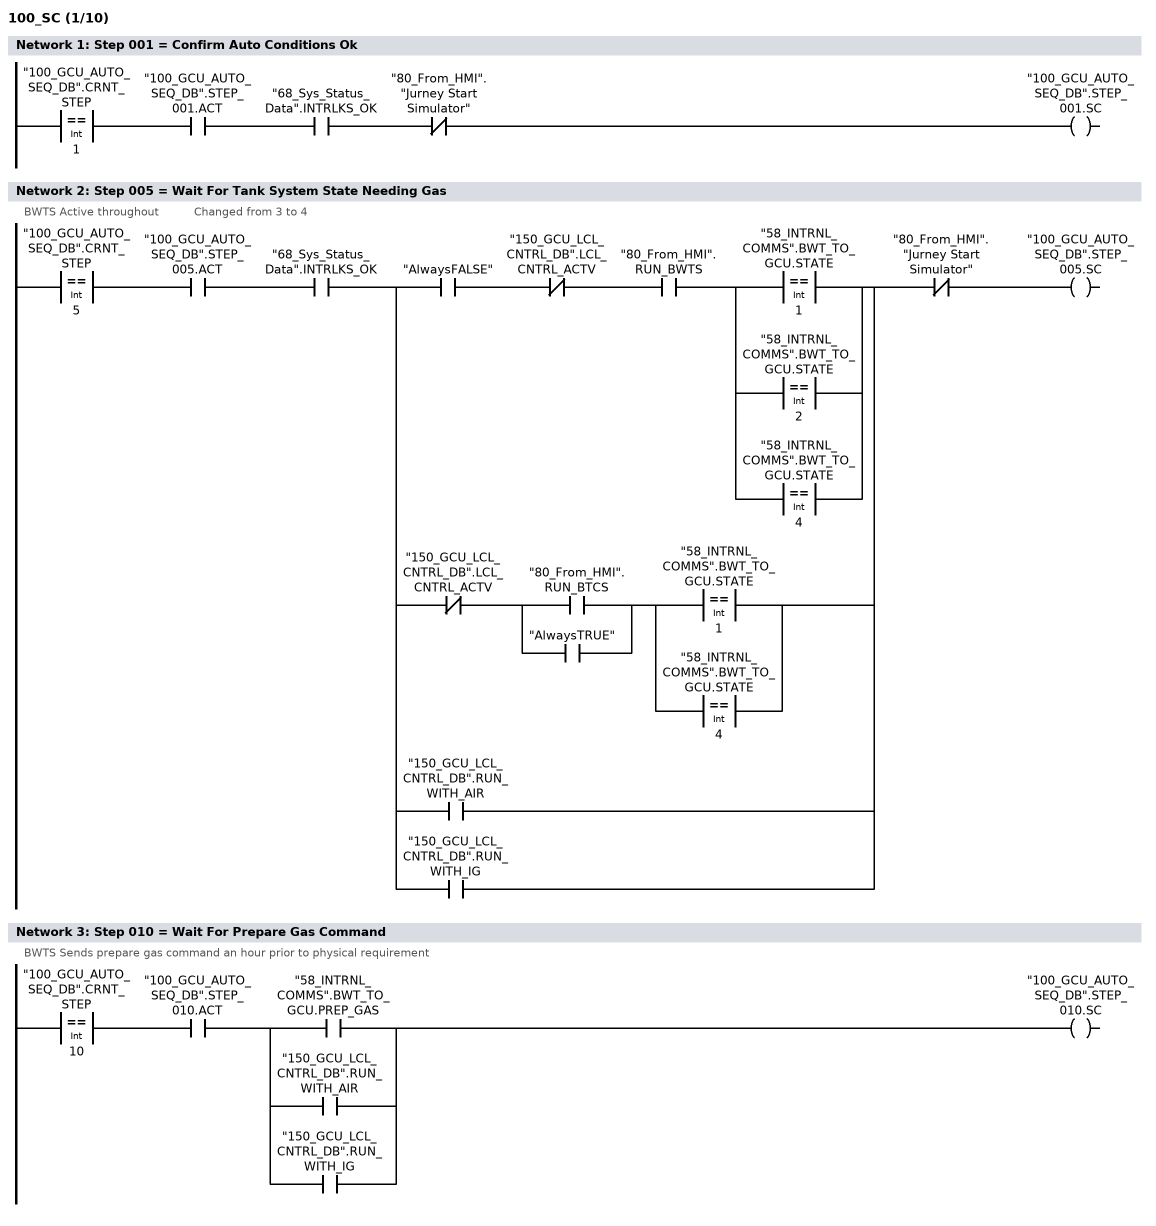
   RUNG wire#powerrail
      { S7_Templates := "SrcType := Int" } EQ_Contact(in1 := "100_GCU_AUTO_SEQ_DB".CRNT_STEP, in2 := 1)
      Contact( "100_GCU_AUTO_SEQ_DB".STEP_001.ACT )
      Contact( "68_Sys_Status_Data".INTRLKS_OK )
      I_Contact( "80_From_HMI"."Jurney Start Simulator" )
      Coil( "100_GCU_AUTO_SEQ_DB".STEP_001.SC )
   END_RUNG
   // the same network as SCL:
   "100_GCU_AUTO_SEQ_DB".STEP_001.SC := ("100_GCU_AUTO_SEQ_DB".CRNT_STEP = 1) AND "100_GCU_AUTO_SEQ_DB".STEP_001.ACT AND "68_Sys_Status_Data".INTRLKS_OK AND NOT "80_From_HMI"."Jurney Start Simulator";
END_REGION

REGION Network 2: Step 005 = Wait For Tank System State Needing Gas
   // BWTS Active throughout          Changed from 3 to 4
   RUNG wire#powerrail
      { S7_Templates := "SrcType := Int" } EQ_Contact(in1 := "100_GCU_AUTO_SEQ_DB".CRNT_STEP, in2 := 5)
      Contact( "100_GCU_AUTO_SEQ_DB".STEP_005.ACT )
      Contact( "68_Sys_Status_Data".INTRLKS_OK )
      wire#w1
      Contact( "AlwaysFALSE" )
      I_Contact( "150_GCU_LCL_CNTRL_DB".LCL_CNTRL_ACTV )
      Contact( "80_From_HMI".RUN_BWTS )
      wire#w2
      { S7_Templates := "SrcType := Int" } EQ_Contact(in1 := "58_INTRNL_COMMS".BWT_TO_GCU.STATE, in2 := 1)
      wire#w3
      I_Contact( "80_From_HMI"."Jurney Start Simulator" )
      Coil( "100_GCU_AUTO_SEQ_DB".STEP_005.SC )
   END_RUNG
   RUNG wire#w2
      { S7_Templates := "SrcType := Int" } EQ_Contact(in1 := "58_INTRNL_COMMS".BWT_TO_GCU.STATE, in2 := 2)
   END_RUNG wire#w3
   RUNG wire#w2
      { S7_Templates := "SrcType := Int" } EQ_Contact(in1 := "58_INTRNL_COMMS".BWT_TO_GCU.STATE, in2 := 4)
   END_RUNG wire#w3
   RUNG wire#w1
      I_Contact( "150_GCU_LCL_CNTRL_DB".LCL_CNTRL_ACTV )
      wire#w4
      Contact( "80_From_HMI".RUN_BTCS )
      wire#w5
      { S7_Templates := "SrcType := Int" } EQ_Contact(in1 := "58_INTRNL_COMMS".BWT_TO_GCU.STATE, in2 := 1)
   END_RUNG wire#w3
   RUNG wire#w4
      Contact( "AlwaysTRUE" )
   END_RUNG wire#w5
   RUNG wire#w5
      { S7_Templates := "SrcType := Int" } EQ_Contact(in1 := "58_INTRNL_COMMS".BWT_TO_GCU.STATE, in2 := 4)
   END_RUNG wire#w3
   RUNG wire#w1
      Contact( "150_GCU_LCL_CNTRL_DB".RUN_WITH_AIR )
   END_RUNG wire#w3
   RUNG wire#w1
      Contact( "150_GCU_LCL_CNTRL_DB".RUN_WITH_IG )
   END_RUNG wire#w3
   // the same network as SCL:
   "100_GCU_AUTO_SEQ_DB".STEP_005.SC := ("100_GCU_AUTO_SEQ_DB".CRNT_STEP = 5) AND "100_GCU_AUTO_SEQ_DB".STEP_005.ACT AND "68_Sys_Status_Data".INTRLKS_OK AND (("AlwaysFALSE" AND NOT "150_GCU_LCL_CNTRL_DB".LCL_CNTRL_ACTV AND "80_From_HMI".RUN_BWTS AND (("58_INTRNL_COMMS".BWT_TO_GCU.STATE = 1) OR ("58_INTRNL_COMMS".BWT_TO_GCU.STATE = 2) OR ("58_INTRNL_COMMS".BWT_TO_GCU.STATE = 4))) OR (NOT "150_GCU_LCL_CNTRL_DB".LCL_CNTRL_ACTV AND ("80_From_HMI".RUN_BTCS OR "AlwaysTRUE") AND (("58_INTRNL_COMMS".BWT_TO_GCU.STATE = 1) OR ("58_INTRNL_COMMS".BWT_TO_GCU.STATE = 4))) OR "150_GCU_LCL_CNTRL_DB".RUN_WITH_AIR OR "150_GCU_LCL_CNTRL_DB".RUN_WITH_IG) AND NOT "80_From_HMI"."Jurney Start Simulator";
END_REGION

REGION Network 3: Step 010 = Wait For Prepare Gas Command
   // BWTS Sends prepare gas command an hour prior to physical requirement
   RUNG wire#powerrail
      { S7_Templates := "SrcType := Int" } EQ_Contact(in1 := "100_GCU_AUTO_SEQ_DB".CRNT_STEP, in2 := 10)
      Contact( "100_GCU_AUTO_SEQ_DB".STEP_010.ACT )
      wire#w1
      Contact( "58_INTRNL_COMMS".BWT_TO_GCU.PREP_GAS )
      wire#w2
      Coil( "100_GCU_AUTO_SEQ_DB".STEP_010.SC )
   END_RUNG
   RUNG wire#w1
      Contact( "150_GCU_LCL_CNTRL_DB".RUN_WITH_AIR )
   END_RUNG wire#w2
   RUNG wire#w1
      Contact( "150_GCU_LCL_CNTRL_DB".RUN_WITH_IG )
   END_RUNG wire#w2
   // the same network as SCL:
   "100_GCU_AUTO_SEQ_DB".STEP_010.SC := ("100_GCU_AUTO_SEQ_DB".CRNT_STEP = 10) AND "100_GCU_AUTO_SEQ_DB".STEP_010.ACT AND ("58_INTRNL_COMMS".BWT_TO_GCU.PREP_GAS OR "150_GCU_LCL_CNTRL_DB".RUN_WITH_AIR OR "150_GCU_LCL_CNTRL_DB".RUN_WITH_IG);
END_REGION

REGION Network 4: Step 020 = Run Command To IGG
   // BWTS Sends prepare gas command an hour prior to physical requirement
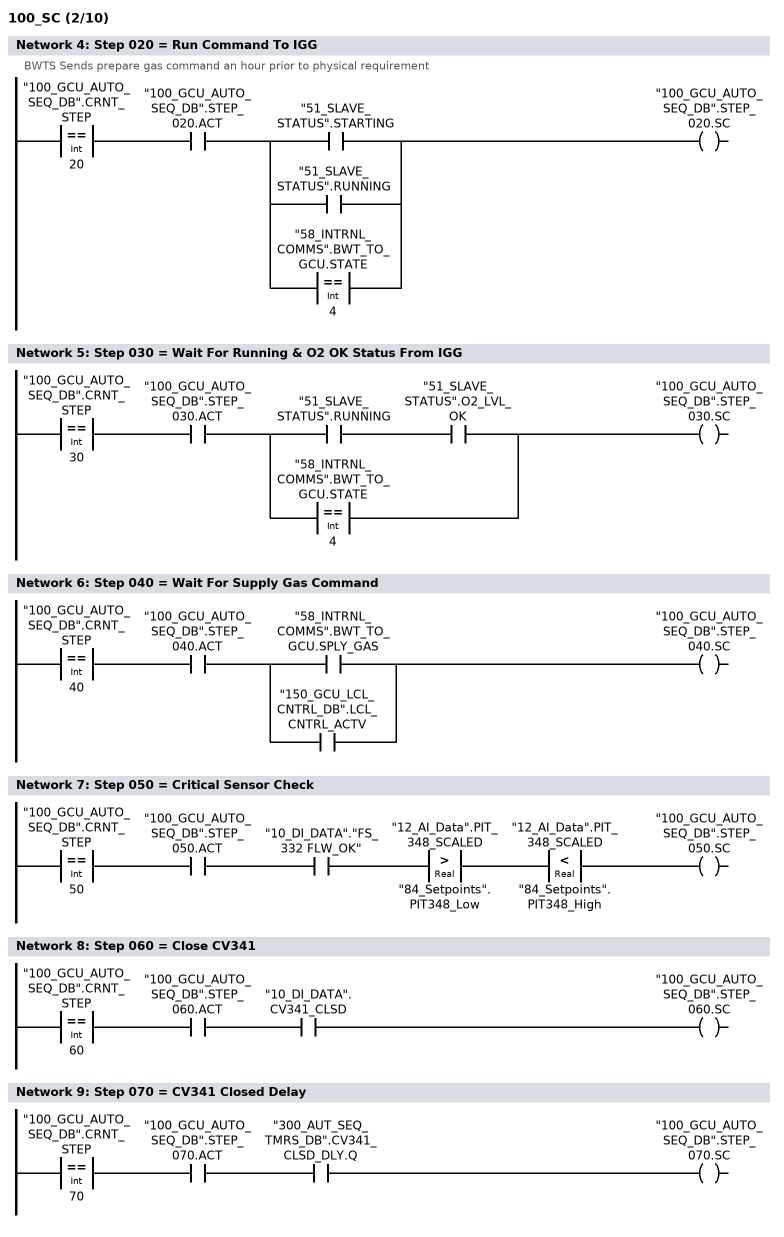
   RUNG wire#powerrail
      { S7_Templates := "SrcType := Int" } EQ_Contact(in1 := "100_GCU_AUTO_SEQ_DB".CRNT_STEP, in2 := 20)
      Contact( "100_GCU_AUTO_SEQ_DB".STEP_020.ACT )
      wire#w1
      Contact( "51_SLAVE_STATUS".STARTING )
      wire#w2
      Coil( "100_GCU_AUTO_SEQ_DB".STEP_020.SC )
   END_RUNG
   RUNG wire#w1
      Contact( "51_SLAVE_STATUS".RUNNING )
   END_RUNG wire#w2
   RUNG wire#w1
      { S7_Templates := "SrcType := Int" } EQ_Contact(in1 := "58_INTRNL_COMMS".BWT_TO_GCU.STATE, in2 := 4)
   END_RUNG wire#w2
   // the same network as SCL:
   "100_GCU_AUTO_SEQ_DB".STEP_020.SC := ("100_GCU_AUTO_SEQ_DB".CRNT_STEP = 20) AND "100_GCU_AUTO_SEQ_DB".STEP_020.ACT AND ("51_SLAVE_STATUS".STARTING OR "51_SLAVE_STATUS".RUNNING OR ("58_INTRNL_COMMS".BWT_TO_GCU.STATE = 4));
END_REGION

REGION Network 5: Step 030 = Wait For Running & O2 OK Status From IGG
   RUNG wire#powerrail
      { S7_Templates := "SrcType := Int" } EQ_Contact(in1 := "100_GCU_AUTO_SEQ_DB".CRNT_STEP, in2 := 30)
      Contact( "100_GCU_AUTO_SEQ_DB".STEP_030.ACT )
      wire#w1
      Contact( "51_SLAVE_STATUS".RUNNING )
      Contact( "51_SLAVE_STATUS".O2_LVL_OK )
      wire#w2
      Coil( "100_GCU_AUTO_SEQ_DB".STEP_030.SC )
   END_RUNG
   RUNG wire#w1
      { S7_Templates := "SrcType := Int" } EQ_Contact(in1 := "58_INTRNL_COMMS".BWT_TO_GCU.STATE, in2 := 4)
   END_RUNG wire#w2
   // the same network as SCL:
   "100_GCU_AUTO_SEQ_DB".STEP_030.SC := ("100_GCU_AUTO_SEQ_DB".CRNT_STEP = 30) AND "100_GCU_AUTO_SEQ_DB".STEP_030.ACT AND (("51_SLAVE_STATUS".RUNNING AND "51_SLAVE_STATUS".O2_LVL_OK) OR ("58_INTRNL_COMMS".BWT_TO_GCU.STATE = 4));
END_REGION

REGION Network 6: Step 040 = Wait For Supply Gas Command
   RUNG wire#powerrail
      { S7_Templates := "SrcType := Int" } EQ_Contact(in1 := "100_GCU_AUTO_SEQ_DB".CRNT_STEP, in2 := 40)
      Contact( "100_GCU_AUTO_SEQ_DB".STEP_040.ACT )
      wire#w1
      Contact( "58_INTRNL_COMMS".BWT_TO_GCU.SPLY_GAS )
      wire#w2
      Coil( "100_GCU_AUTO_SEQ_DB".STEP_040.SC )
   END_RUNG
   RUNG wire#w1
      Contact( "150_GCU_LCL_CNTRL_DB".LCL_CNTRL_ACTV )
   END_RUNG wire#w2
   // the same network as SCL:
   "100_GCU_AUTO_SEQ_DB".STEP_040.SC := ("100_GCU_AUTO_SEQ_DB".CRNT_STEP = 40) AND "100_GCU_AUTO_SEQ_DB".STEP_040.ACT AND ("58_INTRNL_COMMS".BWT_TO_GCU.SPLY_GAS OR "150_GCU_LCL_CNTRL_DB".LCL_CNTRL_ACTV);
END_REGION

REGION Network 7: Step 050 = Critical Sensor Check
   RUNG wire#powerrail
      { S7_Templates := "SrcType := Int" } EQ_Contact(in1 := "100_GCU_AUTO_SEQ_DB".CRNT_STEP, in2 := 50)
      Contact( "100_GCU_AUTO_SEQ_DB".STEP_050.ACT )
      Contact( "10_DI_DATA"."FS_332 FLW_OK" )
      { S7_Templates := "SrcType := Real" } GT_Contact(in1 := "12_AI_Data".PIT_348_SCALED, in2 := "84_Setpoints".PIT348_Low)
      { S7_Templates := "SrcType := Real" } LT_Contact(in1 := "12_AI_Data".PIT_348_SCALED, in2 := "84_Setpoints".PIT348_High)
      Coil( "100_GCU_AUTO_SEQ_DB".STEP_050.SC )
   END_RUNG
   // the same network as SCL:
   "100_GCU_AUTO_SEQ_DB".STEP_050.SC := ("100_GCU_AUTO_SEQ_DB".CRNT_STEP = 50) AND "100_GCU_AUTO_SEQ_DB".STEP_050.ACT AND "10_DI_DATA"."FS_332 FLW_OK" AND ("12_AI_Data".PIT_348_SCALED > "84_Setpoints".PIT348_Low) AND ("12_AI_Data".PIT_348_SCALED < "84_Setpoints".PIT348_High);
END_REGION

REGION Network 8: Step 060 = Close CV341
   RUNG wire#powerrail
      { S7_Templates := "SrcType := Int" } EQ_Contact(in1 := "100_GCU_AUTO_SEQ_DB".CRNT_STEP, in2 := 60)
      Contact( "100_GCU_AUTO_SEQ_DB".STEP_060.ACT )
      Contact( "10_DI_DATA".CV341_CLSD )
      Coil( "100_GCU_AUTO_SEQ_DB".STEP_060.SC )
   END_RUNG
   // the same network as SCL:
   "100_GCU_AUTO_SEQ_DB".STEP_060.SC := ("100_GCU_AUTO_SEQ_DB".CRNT_STEP = 60) AND "100_GCU_AUTO_SEQ_DB".STEP_060.ACT AND "10_DI_DATA".CV341_CLSD;
END_REGION

REGION Network 9: Step 070 = CV341 Closed Delay
   RUNG wire#powerrail
      { S7_Templates := "SrcType := Int" } EQ_Contact(in1 := "100_GCU_AUTO_SEQ_DB".CRNT_STEP, in2 := 70)
      Contact( "100_GCU_AUTO_SEQ_DB".STEP_070.ACT )
      Contact( "300_AUT_SEQ_TMRS_DB".CV341_CLSD_DLY.Q )
      Coil( "100_GCU_AUTO_SEQ_DB".STEP_070.SC )
   END_RUNG
   // the same network as SCL:
   "100_GCU_AUTO_SEQ_DB".STEP_070.SC := ("100_GCU_AUTO_SEQ_DB".CRNT_STEP = 70) AND "100_GCU_AUTO_SEQ_DB".STEP_070.ACT AND "300_AUT_SEQ_TMRS_DB".CV341_CLSD_DLY.Q;
END_REGION

REGION Network 10: Step 080 = Amend Setpoints
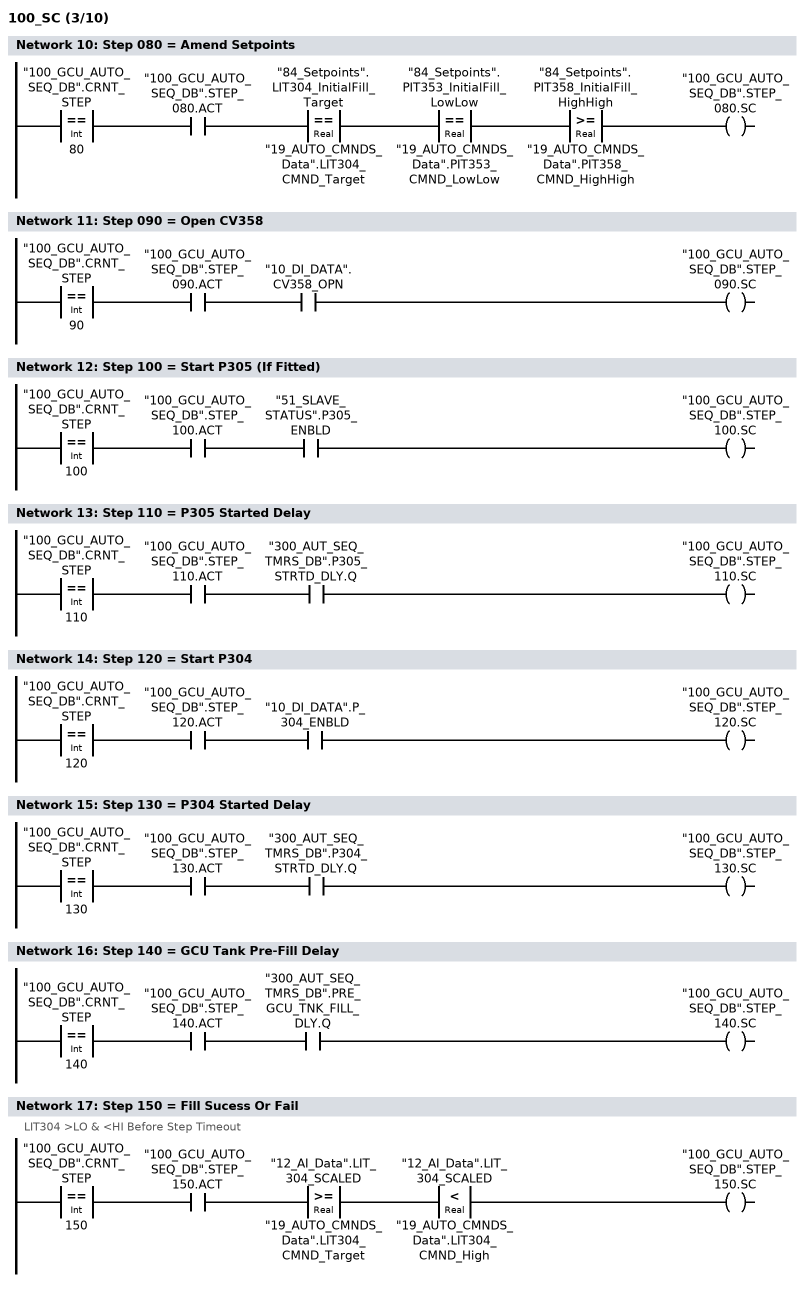
   RUNG wire#powerrail
      { S7_Templates := "SrcType := Int" } EQ_Contact(in1 := "100_GCU_AUTO_SEQ_DB".CRNT_STEP, in2 := 80)
      Contact( "100_GCU_AUTO_SEQ_DB".STEP_080.ACT )
      { S7_Templates := "SrcType := Real" } EQ_Contact(in1 := "84_Setpoints".LIT304_InitialFill_Target, in2 := "19_AUTO_CMNDS_Data".LIT304_CMND_Target)
      { S7_Templates := "SrcType := Real" } EQ_Contact(in1 := "84_Setpoints".PIT353_InitialFill_LowLow, in2 := "19_AUTO_CMNDS_Data".PIT353_CMND_LowLow)
      { S7_Templates := "SrcType := Real" } GE_Contact(in1 := "84_Setpoints".PIT358_InitialFill_HighHigh, in2 := "19_AUTO_CMNDS_Data".PIT358_CMND_HighHigh)
      Coil( "100_GCU_AUTO_SEQ_DB".STEP_080.SC )
   END_RUNG
   // the same network as SCL:
   "100_GCU_AUTO_SEQ_DB".STEP_080.SC := ("100_GCU_AUTO_SEQ_DB".CRNT_STEP = 80) AND "100_GCU_AUTO_SEQ_DB".STEP_080.ACT AND ("84_Setpoints".LIT304_InitialFill_Target = "19_AUTO_CMNDS_Data".LIT304_CMND_Target) AND ("84_Setpoints".PIT353_InitialFill_LowLow = "19_AUTO_CMNDS_Data".PIT353_CMND_LowLow) AND ("84_Setpoints".PIT358_InitialFill_HighHigh >= "19_AUTO_CMNDS_Data".PIT358_CMND_HighHigh);
END_REGION

REGION Network 11: Step 090 = Open CV358
   RUNG wire#powerrail
      { S7_Templates := "SrcType := Int" } EQ_Contact(in1 := "100_GCU_AUTO_SEQ_DB".CRNT_STEP, in2 := 90)
      Contact( "100_GCU_AUTO_SEQ_DB".STEP_090.ACT )
      Contact( "10_DI_DATA".CV358_OPN )
      Coil( "100_GCU_AUTO_SEQ_DB".STEP_090.SC )
   END_RUNG
   // the same network as SCL:
   "100_GCU_AUTO_SEQ_DB".STEP_090.SC := ("100_GCU_AUTO_SEQ_DB".CRNT_STEP = 90) AND "100_GCU_AUTO_SEQ_DB".STEP_090.ACT AND "10_DI_DATA".CV358_OPN;
END_REGION

REGION Network 12: Step 100 = Start P305 (If Fitted)
   RUNG wire#powerrail
      { S7_Templates := "SrcType := Int" } EQ_Contact(in1 := "100_GCU_AUTO_SEQ_DB".CRNT_STEP, in2 := 100)
      Contact( "100_GCU_AUTO_SEQ_DB".STEP_100.ACT )
      Contact( "51_SLAVE_STATUS".P305_ENBLD )
      Coil( "100_GCU_AUTO_SEQ_DB".STEP_100.SC )
   END_RUNG
   // the same network as SCL:
   "100_GCU_AUTO_SEQ_DB".STEP_100.SC := ("100_GCU_AUTO_SEQ_DB".CRNT_STEP = 100) AND "100_GCU_AUTO_SEQ_DB".STEP_100.ACT AND "51_SLAVE_STATUS".P305_ENBLD;
END_REGION

REGION Network 13: Step 110 = P305 Started Delay
   RUNG wire#powerrail
      { S7_Templates := "SrcType := Int" } EQ_Contact(in1 := "100_GCU_AUTO_SEQ_DB".CRNT_STEP, in2 := 110)
      Contact( "100_GCU_AUTO_SEQ_DB".STEP_110.ACT )
      Contact( "300_AUT_SEQ_TMRS_DB".P305_STRTD_DLY.Q )
      Coil( "100_GCU_AUTO_SEQ_DB".STEP_110.SC )
   END_RUNG
   // the same network as SCL:
   "100_GCU_AUTO_SEQ_DB".STEP_110.SC := ("100_GCU_AUTO_SEQ_DB".CRNT_STEP = 110) AND "100_GCU_AUTO_SEQ_DB".STEP_110.ACT AND "300_AUT_SEQ_TMRS_DB".P305_STRTD_DLY.Q;
END_REGION

REGION Network 14: Step 120 = Start P304
   RUNG wire#powerrail
      { S7_Templates := "SrcType := Int" } EQ_Contact(in1 := "100_GCU_AUTO_SEQ_DB".CRNT_STEP, in2 := 120)
      Contact( "100_GCU_AUTO_SEQ_DB".STEP_120.ACT )
      Contact( "10_DI_DATA".P_304_ENBLD )
      Coil( "100_GCU_AUTO_SEQ_DB".STEP_120.SC )
   END_RUNG
   // the same network as SCL:
   "100_GCU_AUTO_SEQ_DB".STEP_120.SC := ("100_GCU_AUTO_SEQ_DB".CRNT_STEP = 120) AND "100_GCU_AUTO_SEQ_DB".STEP_120.ACT AND "10_DI_DATA".P_304_ENBLD;
END_REGION

REGION Network 15: Step 130 = P304 Started Delay
   RUNG wire#powerrail
      { S7_Templates := "SrcType := Int" } EQ_Contact(in1 := "100_GCU_AUTO_SEQ_DB".CRNT_STEP, in2 := 130)
      Contact( "100_GCU_AUTO_SEQ_DB".STEP_130.ACT )
      Contact( "300_AUT_SEQ_TMRS_DB".P304_STRTD_DLY.Q )
      Coil( "100_GCU_AUTO_SEQ_DB".STEP_130.SC )
   END_RUNG
   // the same network as SCL:
   "100_GCU_AUTO_SEQ_DB".STEP_130.SC := ("100_GCU_AUTO_SEQ_DB".CRNT_STEP = 130) AND "100_GCU_AUTO_SEQ_DB".STEP_130.ACT AND "300_AUT_SEQ_TMRS_DB".P304_STRTD_DLY.Q;
END_REGION

REGION Network 16: Step 140 = GCU Tank Pre-Fill Delay
   RUNG wire#powerrail
      { S7_Templates := "SrcType := Int" } EQ_Contact(in1 := "100_GCU_AUTO_SEQ_DB".CRNT_STEP, in2 := 140)
      Contact( "100_GCU_AUTO_SEQ_DB".STEP_140.ACT )
      Contact( "300_AUT_SEQ_TMRS_DB".PRE_GCU_TNK_FILL_DLY.Q )
      Coil( "100_GCU_AUTO_SEQ_DB".STEP_140.SC )
   END_RUNG
   // the same network as SCL:
   "100_GCU_AUTO_SEQ_DB".STEP_140.SC := ("100_GCU_AUTO_SEQ_DB".CRNT_STEP = 140) AND "100_GCU_AUTO_SEQ_DB".STEP_140.ACT AND "300_AUT_SEQ_TMRS_DB".PRE_GCU_TNK_FILL_DLY.Q;
END_REGION

REGION Network 17: Step 150 = Fill Sucess Or Fail
   // LIT304 >LO & <HI Before Step Timeout
   RUNG wire#powerrail
      { S7_Templates := "SrcType := Int" } EQ_Contact(in1 := "100_GCU_AUTO_SEQ_DB".CRNT_STEP, in2 := 150)
      Contact( "100_GCU_AUTO_SEQ_DB".STEP_150.ACT )
      { S7_Templates := "SrcType := Real" } GE_Contact(in1 := "12_AI_Data".LIT_304_SCALED, in2 := "19_AUTO_CMNDS_Data".LIT304_CMND_Target)
      { S7_Templates := "SrcType := Real" } LT_Contact(in1 := "12_AI_Data".LIT_304_SCALED, in2 := "19_AUTO_CMNDS_Data".LIT304_CMND_High)
      Coil( "100_GCU_AUTO_SEQ_DB".STEP_150.SC )
   END_RUNG
   // the same network as SCL:
   "100_GCU_AUTO_SEQ_DB".STEP_150.SC := ("100_GCU_AUTO_SEQ_DB".CRNT_STEP = 150) AND "100_GCU_AUTO_SEQ_DB".STEP_150.ACT AND ("12_AI_Data".LIT_304_SCALED >= "19_AUTO_CMNDS_Data".LIT304_CMND_Target) AND ("12_AI_Data".LIT_304_SCALED < "19_AUTO_CMNDS_Data".LIT304_CMND_High);
END_REGION

REGION Network 18: Step 160 = Stop P304
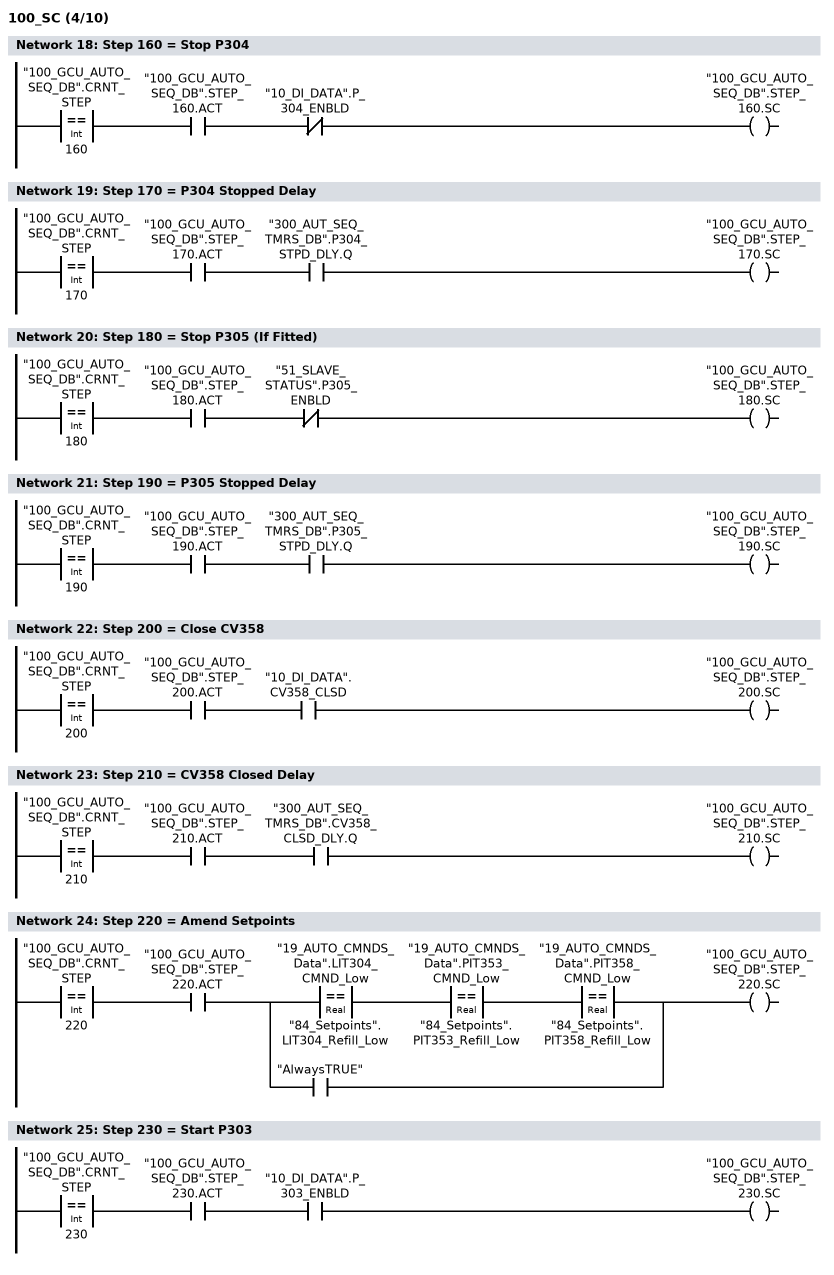
   RUNG wire#powerrail
      { S7_Templates := "SrcType := Int" } EQ_Contact(in1 := "100_GCU_AUTO_SEQ_DB".CRNT_STEP, in2 := 160)
      Contact( "100_GCU_AUTO_SEQ_DB".STEP_160.ACT )
      I_Contact( "10_DI_DATA".P_304_ENBLD )
      Coil( "100_GCU_AUTO_SEQ_DB".STEP_160.SC )
   END_RUNG
   // the same network as SCL:
   "100_GCU_AUTO_SEQ_DB".STEP_160.SC := ("100_GCU_AUTO_SEQ_DB".CRNT_STEP = 160) AND "100_GCU_AUTO_SEQ_DB".STEP_160.ACT AND NOT "10_DI_DATA".P_304_ENBLD;
END_REGION
